// TIA Portal project "Industry 4.0_Plant_Logic" (V16)

(* hardware
DEVICE "S7-1200 station_1"  S7-1200 Station
   slot 0: "Rack_0"  S7-1200 Rack  Rack  V1.0
   slot 1: "S7_1212"  CPU 1212C AC/DC/Rly  6ES7 212-1BE40-0XB0  V4.4
   slot 2: "AQ 2x14BIT_1"  SM 1232 AQ2  6ES7 232-4HB32-0XB0  V2.1
DEVICE "HMI_1"  KTP700 Basic PN
   slot 0: "HMI_1"  KTP700 Basic PN  6AV2 123-2GB03-0AX0  15.1.0.0
   slot 1: "HMI_RT_1"  KTP700 Basic PN  6AV2 123-2GB03-0AX0  15.1.0.0
   slot 5: "HMI_1.IE_CP_1"  PROFINET Interface  15.0.1.0
      slot 1: "PROFINET Interface_1"  PROFINET Interface
         slot 1: "Port_1"  Port
*)

// ===== PLC "S7_1212"  CPU 1212C AC/DC/Rly =====

VAR_GLOBAL   // PLC tag table "Default tag table"
   "FIC_B102" AT %IW64 : Int;   // Flow meter(0 - 27648)
   "LIC_B101" AT %IW66 : Int;   // Tank02 Level meter(0 - 27648)
   "PS1_RFID_Station" AT %I0.0 : Bool;   // PS-Proximity Switch
   "PS2_Filling_Station" AT %I0.1 : Bool;
   "PS3_Quality_Station" AT %I0.2 : Bool;
   "PS4_End_of_Conveyor" AT %I0.3 : Bool;
   "T01_Low_Level" AT %I0.4 : Bool;   // Proximity sensor measuring Low level of Tank01
   "T01_High_Level" AT %I0.5 : Bool;   // Proximity sensor measuring High level of Tank01
   "T01_Outlet" AT %Q0.1 : Bool;   // Tank01 Output Solenoid Valve
   "T02_Outlet" AT %Q0.2 : Bool;   // Tank02 Output Solenoid Valve
   "Outlet_Pump_Motor" AT %Q0.3 : Bool;   // Pump Motor
   "Conveyor_Motor" AT %Q0.0 : Bool;
   "NTRG_06" AT %M5.5 : Bool;
   "NTRG_09" AT %M5.6 : Bool;
   "NTRG_099" AT %M5.7 : Bool;
   "PTRG10" AT %M6.0 : Bool;
   "PTRIG999" AT %M6.1 : Bool;
   "PTRIG998" AT %M6.2 : Bool;
   "PTRIG888" AT %M6.3 : Bool;
   "ptrig141" AT %M6.4 : Bool;
   "ptrig142" AT %M6.5 : Bool;
   "ptrig143" AT %M6.6 : Bool;
   "Ptrig241" AT %M6.7 : Bool;
   "reset__bottle_animation_timer" AT %M7.0 : Bool;
   "motor_running_time" AT %MD8 : Time;
   "ntrig555" AT %M7.1 : Bool;
   "Total Bottle filled" AT %MW8 : Int;
   "abc" AT %QW98 : Int;
   "Static_1" AT %MW12 : Int;
   "Static_1(1)" AT %MW14 : Int;
   "Static_1(2)" AT %MW16 : Int;
   "i" AT %MW18 : Int;
   "ONS_1" AT %M7.2 : Bool;
END_VAR

VAR_GLOBAL   // PLC tag table "P_N_TRIG"
   "PTRIG1" AT %M0.0 : Bool;
   "PTRIG2" AT %M0.1 : Bool;
   "PTRIG3" AT %M0.2 : Bool;
   "PTRIG4" AT %M0.3 : Bool;
   "PTRIG5" AT %M0.4 : Bool;
   "PTRIG6" AT %M0.5 : Bool;
   "PTRIG7" AT %M0.6 : Bool;
   "PTRIG8" AT %M0.7 : Bool;
   "PTRIG9" AT %M1.0 : Bool;
   "PTRIG10" AT %M1.1 : Bool;
   "PTRIG11" AT %M1.2 : Bool;
   "PTRIG12" AT %M1.3 : Bool;
   "PTRIG13" AT %M1.4 : Bool;
   "PTRIG14" AT %M1.5 : Bool;
   "PTRIG15" AT %M1.6 : Bool;
   "PTRIG16" AT %M1.7 : Bool;
   "PTRIG17" AT %M2.0 : Bool;
   "PTRIG18" AT %M2.1 : Bool;
   "PTRIG19" AT %M2.2 : Bool;
   "PTRIG20" AT %M2.3 : Bool;
   "PTRIG21" AT %M2.4 : Bool;
   "PTRIG22" AT %M2.5 : Bool;
   "PTRIG23" AT %M2.6 : Bool;
   "NTRIG1" AT %M2.7 : Bool;
   "NTRIG2" AT %M3.0 : Bool;
   "NTRIG3" AT %M3.1 : Bool;
   "NTRIG4" AT %M3.2 : Bool;
   "NTRIG5" AT %M3.3 : Bool;
   "NTRIG6" AT %M3.4 : Bool;
   "NTRIG7" AT %M3.5 : Bool;
   "NTRIG8" AT %M3.6 : Bool;
   "NTRIG9" AT %M3.7 : Bool;
   "NTRIG10" AT %M4.0 : Bool;
   "NTRIG11" AT %M4.1 : Bool;
   "NTRIG12" AT %M4.2 : Bool;
   "NTRIG13" AT %M4.3 : Bool;
   "NTRIG14" AT %M4.4 : Bool;
   "NTRIG15" AT %M4.5 : Bool;
   "NTRIG16" AT %M4.6 : Bool;
   "NTRIG17" AT %M4.7 : Bool;
   "NTRIG18" AT %M5.0 : Bool;
   "NTRIG19" AT %M5.1 : Bool;
   "NTRIG20" AT %M5.2 : Bool;
   "PTRIG24" AT %M5.3 : Bool;
   "PTRIG25" AT %M5.4 : Bool;
END_VAR

DATA_BLOCK "Global_DB"   // DB1
{ S7_Optimized_Access := 'TRUE' }
VERSION : 0.1
   VAR
      Input : Struct   // Values from input devices
         FIC_B102 : Int;   // Flow in (0-27648) range
         LIC_B101 : Int;   // Level in (0-27648) range
         PS1_RFID_Station : Bool;   // Proximity sensor at RFID station
         PS2_Filling_Station : Bool;   // Proximity sensor at Filling station
         PS3_Quality_Station : Bool;   // Proximity sensor at Quality Station
         PS4_End_of_Conveyor : Bool;   // Proximity sensor at End of the conveyor
         T01_Low_Level : Bool;   // Tank01 Low level detection sensor
         T01_High_Level : Bool;   // Tank01 High level detection sensor
      END_STRUCT;
      Output : Struct   // Values to Output devices
         T01_Outlet : Bool;   // Tank01 Outlet Solenoid Valve
         T02_Outlet : Bool;   // Tank02 Outlet Solenoid Valve
         Outlet_Pump_Motor : Bool;   // To tigger Pump motor relay
         Conveyor_Motor : Bool;   // To tigger Conveyor motor relay
         T01_Inlet : Bool;   // Tank01 Inlet Solenoid Valve(Not implemented)
         T02_Inlet : Bool;   // Tank02 Inlet Solenoid Valve(Not implemented)
      END_STRUCT;
      Other_Parameters : Struct   // Scalled and middle Variables
         Liquid_A_Filled : Bool;   // Liquid_A_filled flag activated when intended amount of Liquid A is filled
         Add_Done : Bool;
         Liquid_B_Filled : Bool;   // Liquid_B_filled flag activated when intended amount of Liquid B is filled
         Flow_ml_per_sec : Real;   // Scalled flow meter reading (0-250mL/sec)
         LiquidA_in_Bottle_ml : Real;
         LiquidB_in_Bottle_ml : Real;
         T02_Level_in_L : Real;   // Scalled level meter reading (0-10L)
         T02_High_Level_Limit : Real;
         T02_Low_Level_Limit : Real;
         Alarm_Reset : Bool;   // to reset all active alarms
         operation_cycle_time : Time;   // Time taken for the filling of one bottle
         index : Int := 1;
      END_STRUCT;
      Error : Struct
         Alarm : Word;
      END_STRUCT;
      Master_Commands : Struct
         operation_finished : Bool;
         operation_begin : Bool;
         Order_Variables : Struct   // Online Order parameter
            "Total Bottle filled" : Int;
            Order_ID : UInt;
            Quantity : UInt := 0;   // Quanity of bottle to be filled in pesent order
            Liquid_A_pct : Int := 0;   // data from RFID tags or Order
            Liquid_B_pct : Int;   // datafrom RFID tags or Order
            Order_received : Bool;   // Activated when new order is received.
            Bottle_Count : Int := 1;   // Total Bottle filled
            Order_completed : Bool;   // Order completion flag(After filling all bottle)
         END_STRUCT;
      END_STRUCT;
      SCADA : Struct   // SCADA animation tags
         motor_running_time : Time;   // To display bottle moving on the conveyor based on the running time of conveyor
      END_STRUCT;
      Flow : Real;
      Motor_Output_PCT : Int;
      Production_Data : Struct   // Unit ml
         Total_Liquid_in_Bottle : Array[1..5] of Real;
         LiquidA_in_Bottle : Array[1..5] of Real;
         operation_cycles : Array[1..5] of Time;
         LiquidB_in_Bottle : Array[1..5] of Real;
         current_cycle : Int := 1;
      END_STRUCT;
      Array_Voltage : Array[0..999] of Real;
      Voltage_Timer : Bool;
      "Locking bits" : Struct
         Starting_station_bit : Bool;
         Filling_station_bit : Bool;
         Quality_station_bit : Bool;
         End_station_bit : Bool;
      END_STRUCT;
   END_VAR
BEGIN
END_DATA_BLOCK

// folder: Function Blocks

DATA_BLOCK "Re-filling_Logic_DB"   // DB2
{ S7_Optimized_Access := 'TRUE' }
VERSION : 0.1
// stored: InstanceOfName Re-filling_Logic
"Re-filling_Logic"
BEGIN
END_DATA_BLOCK

DATA_BLOCK "Filling_Logic_DB"   // DB4
{ S7_Optimized_Access := 'TRUE' }
VERSION : 0.1
// stored: InstanceOfName Filling_Logic
"Filling_Logic"
BEGIN
END_DATA_BLOCK

DATA_BLOCK "Filling_Logic_DB_1"   // DB5
{ S7_Optimized_Access := 'TRUE' }
VERSION : 0.1
// stored: InstanceOfName Filling_Logic
"Filling_Logic"
BEGIN
END_DATA_BLOCK

DATA_BLOCK "Alarm_Logic_DB"   // DB7
{ S7_Optimized_Access := 'TRUE' }
VERSION : 0.1
// stored: InstanceOfName Alarm_Logic
"Alarm_Logic"
BEGIN
END_DATA_BLOCK

DATA_BLOCK "Tank1_DB"   // DB9
{ S7_Optimized_Access := 'TRUE' }
VERSION : 0.1
// stored: InstanceOfName Tank1
"Tank1"
BEGIN
END_DATA_BLOCK

DATA_BLOCK "Tank2_DB"   // DB10
{ S7_Optimized_Access := 'TRUE' }
VERSION : 0.1
// stored: InstanceOfName Tank2
"Tank2"
BEGIN
END_DATA_BLOCK

DATA_BLOCK "ProductionData_Reset_DB"   // DB13
{ S7_Optimized_Access := 'TRUE' }
VERSION : 0.1
// stored: InstanceOfName ProductionData_Reset
"ProductionData_Reset"
BEGIN
END_DATA_BLOCK

DATA_BLOCK "Operation_cycle_DB"   // DB15
{ S7_Optimized_Access := 'TRUE' }
VERSION : 0.1
// stored: InstanceOfName Operation_cycle
"Operation_cycle"
BEGIN
END_DATA_BLOCK

DATA_BLOCK "Reseting_order_DB"   // DB18
{ S7_Optimized_Access := 'TRUE' }
VERSION : 0.1
// stored: InstanceOfName Reseting_order
"Reseting_order"
BEGIN
END_DATA_BLOCK

DATA_BLOCK "Array_Voltage_Logic_DB_1"   // DB25
{ S7_Optimized_Access := 'TRUE' }
VERSION : 0.1
// stored: InstanceOfName Array_Voltage_Logic
"Array_Voltage_Logic"
BEGIN
END_DATA_BLOCK

// folder: System blocks/Program resources

DATA_BLOCK "IEC_Timer_6_DB_1"   // DB3
{ S7_Optimized_Access := 'TRUE' }
AUTHOR : Simatic
FAMILY : IEC
NAME : IEC_TMR
VERSION : 1.0
// stored: InstanceOfName IEC_TIMER
"IEC_TIMER"
BEGIN
END_DATA_BLOCK

DATA_BLOCK "IEC_Timer_0_DB_1"   // DB6
{ S7_Optimized_Access := 'TRUE' }
AUTHOR : Simatic
FAMILY : IEC
NAME : IEC_TMR
VERSION : 1.0
// stored: InstanceOfName IEC_TIMER
"IEC_TIMER"
BEGIN
END_DATA_BLOCK

DATA_BLOCK "IEC_Timer_0_DB_999"   // DB8
{ S7_Optimized_Access := 'TRUE' }
AUTHOR : Simatic
FAMILY : IEC
NAME : IEC_TMR
VERSION : 1.0
// stored: InstanceOfName IEC_TIMER
"IEC_TIMER"
BEGIN
END_DATA_BLOCK

DATA_BLOCK "IEC_Timer_0_DB_7"   // DB11
{ S7_Optimized_Access := 'TRUE' }
AUTHOR : Simatic
FAMILY : IEC
NAME : IEC_TMR
VERSION : 1.0
// stored: InstanceOfName IEC_TIMER
"IEC_TIMER"
BEGIN
END_DATA_BLOCK

DATA_BLOCK "IEC_Counter_0_DB"   // DB12
{ S7_Optimized_Access := 'TRUE' }
AUTHOR : Simatic
FAMILY : IEC
NAME : CNTR
VERSION : 1.0
// stored: InstanceOfName IEC_COUNTER
"IEC_COUNTER"
BEGIN
END_DATA_BLOCK

DATA_BLOCK "Cycle_time"   // DB14
{ S7_Optimized_Access := 'TRUE' }
AUTHOR : Simatic
FAMILY : IEC
NAME : IEC_TMR
VERSION : 1.0
// stored: InstanceOfName IEC_TIMER
"IEC_TIMER"
BEGIN
END_DATA_BLOCK

DATA_BLOCK "IEC_Timer_655"   // DB16
{ S7_Optimized_Access := 'TRUE' }
AUTHOR : Simatic
FAMILY : IEC
NAME : IEC_TMR
VERSION : 1.0
// stored: InstanceOfName IEC_TIMER
"IEC_TIMER"
BEGIN
END_DATA_BLOCK

DATA_BLOCK "Waiting time"   // DB20
{ S7_Optimized_Access := 'TRUE' }
AUTHOR : Simatic
FAMILY : IEC
NAME : IEC_TMR
VERSION : 1.0
// stored: InstanceOfName IEC_TIMER
"IEC_TIMER"
BEGIN
END_DATA_BLOCK

// folder: (top level)

ORGANIZATION_BLOCK "Main"   // OB1, LAD, ProgramCycle
TITLE = "Main Program Sweep (Cycle)"
{ S7_Optimized_Access := 'TRUE' }
VERSION : 0.1
   VAR_INPUT
      Initial_Call : Bool;   // Initial call of this OB
      Remanence : Bool;   // =True, if remanent data are available
   END_VAR
   VAR_TEMP   // added for the SCL form of the ladder/FBD networks
      _w1 : Bool;
      _w2 : Bool;
   END_VAR
BEGIN

REGION Network 1: Tank 1 and Tank 2 re-filling Logic
   // 1."Re-filling_logic" block is logic block to refill liquid in tanks based on their levels(Hardware not present yet)
   // 2."Operation_cycle" block to measure the time of bottle filling which starts from picking bottle till bottle placed.
   // 3."Reading" Mapping from Physical address to Global_DB (for input devices)
   // 4."Writing" Mapping from Global_DB to Physical address(for output devices)
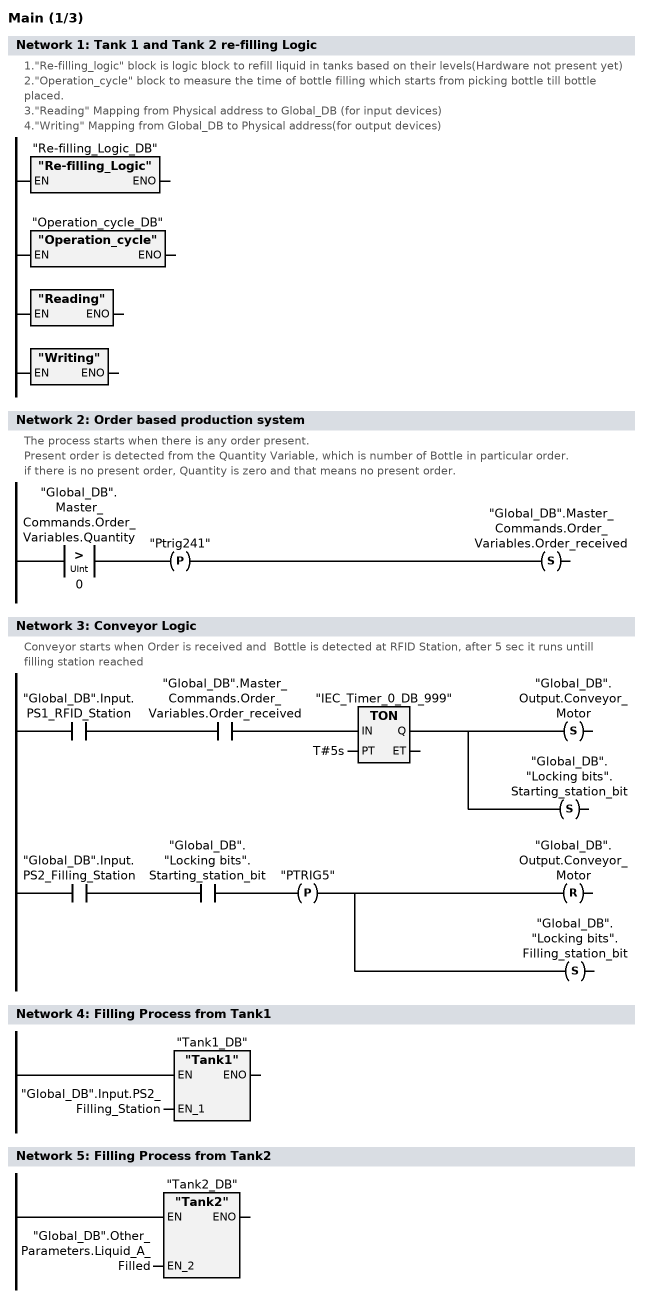
   RUNG wire#powerrail
      "Re-filling_Logic_DB"()
   END_RUNG
   RUNG wire#powerrail
      "Operation_cycle_DB"()
   END_RUNG
   RUNG wire#powerrail
      "Reading"()
   END_RUNG
   RUNG wire#powerrail
      "Writing"()
   END_RUNG
   // the same network as SCL:
   "Re-filling_Logic_DB"();   // "Re-filling_Logic"
   "Operation_cycle_DB"();   // "Operation_cycle"
   "Reading"();
   "Writing"();
END_REGION

REGION Network 2: Order based production system
   // The process starts when there is any order present.
   // Present order is detected from the Quantity Variable, which is number of Bottle in particular order.
   // if there is no present order, Quantity is zero and that means no present order.
   RUNG wire#powerrail
      { S7_Templates := "SrcType := UInt" } GT_Contact(in1 := "Global_DB".Master_Commands.Order_Variables.Quantity, in2 := 0)
      P_Trig( "Ptrig241" )
      S_Coil( "Global_DB".Master_Commands.Order_Variables.Order_received )
   END_RUNG
   // the same network as SCL:
   #_w1 := "Global_DB".Master_Commands.Order_Variables.Quantity > 0;
   #_w2 := #_w1 AND NOT "Ptrig241";   // rising edge
   "Ptrig241" := #_w1;
   IF #_w2 THEN "Global_DB".Master_Commands.Order_Variables.Order_received := TRUE; END_IF;
END_REGION

REGION Network 3: Conveyor Logic
   // Conveyor starts when Order is received and  Bottle is detected at RFID Station, after 5 sec it runs untill filling station reached
   "IEC_Timer_0_DB_999".TON(IN := "Global_DB".Input.PS1_RFID_Station AND "Global_DB".Master_Commands.Order_Variables.Order_received,
                           PT := T#5s);
   IF "IEC_Timer_0_DB_999".Q THEN
       "Global_DB".Output.Conveyor_Motor := TRUE;
       "Global_DB"."Locking bits".Starting_station_bit := TRUE;
   END_IF;
   #_w1 := "Global_DB".Input.PS2_Filling_Station AND "Global_DB"."Locking bits".Starting_station_bit;
   #_w2 := #_w1 AND NOT "PTRIG5";   // rising edge
   "PTRIG5" := #_w1;
   IF #_w2 THEN
       "Global_DB".Output.Conveyor_Motor := FALSE;
       "Global_DB"."Locking bits".Filling_station_bit := TRUE;
   END_IF;
END_REGION

REGION Network 4: Filling Process from Tank1
   RUNG wire#powerrail
      "Tank1_DB"(EN_1 := "Global_DB".Input.PS2_Filling_Station)
   END_RUNG
   // the same network as SCL:
   "Tank1_DB"(EN_1 := "Global_DB".Input.PS2_Filling_Station);   // "Tank1"
END_REGION

REGION Network 5: Filling Process from Tank2
   RUNG wire#powerrail
      "Tank2_DB"(EN_2 := "Global_DB".Other_Parameters.Liquid_A_Filled)
   END_RUNG
   // the same network as SCL:
   "Tank2_DB"(EN_2 := "Global_DB".Other_Parameters.Liquid_A_Filled);   // "Tank2"
END_REGION

REGION Network 6: Store data in database for records
   // after filling the liquid from both tanks, ADD block adds the value of filled amount of Liquid A nad Liquid B in the bottle to keep record of total liquid filled in particular bottle.
   // 
   // then bottle number is incremented.
   // 
   // Values reset for next cycle.
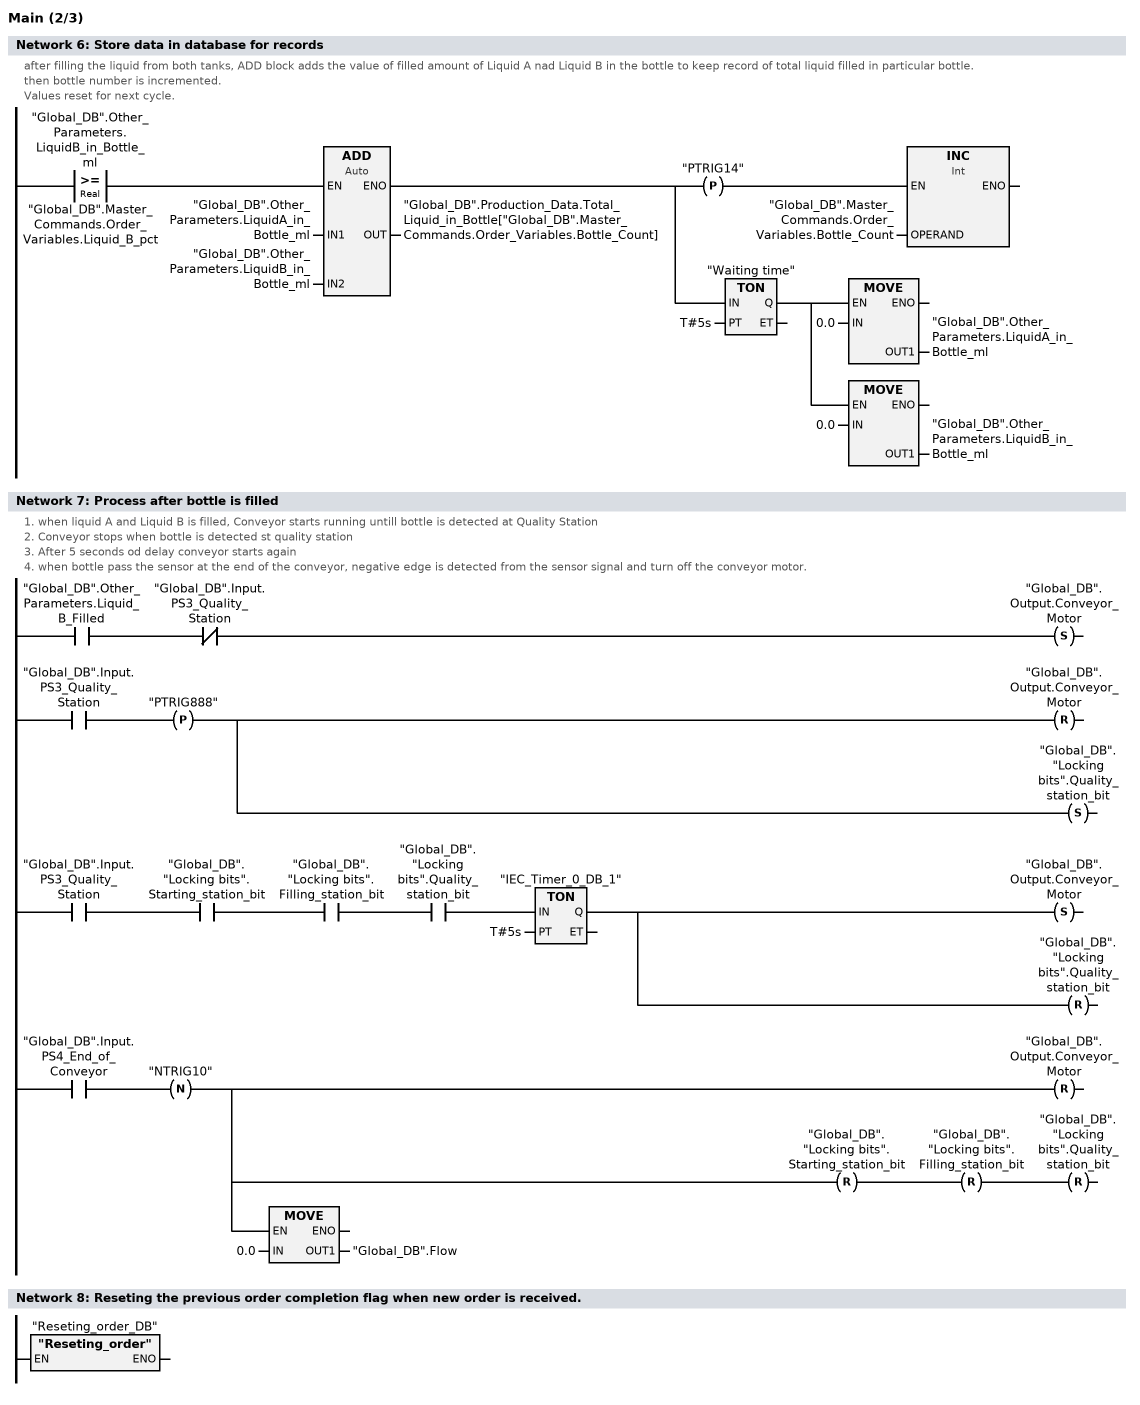
   #_w1 := "Global_DB".Other_Parameters.LiquidB_in_Bottle_ml >= "Global_DB".Master_Commands.Order_Variables.Liquid_B_pct;
   IF #_w1 THEN
       "Global_DB".Production_Data.Total_Liquid_in_Bottle["Global_DB".Master_Commands.Order_Variables.Bottle_Count] := "Global_DB".Other_Parameters.LiquidA_in_Bottle_ml + "Global_DB".Other_Parameters.LiquidB_in_Bottle_ml;
   END_IF;
   #_w2 := #_w1 AND NOT "PTRIG14";   // rising edge
   "PTRIG14" := #_w1;
   IF #_w2 THEN
       "Global_DB".Master_Commands.Order_Variables.Bottle_Count := "Global_DB".Master_Commands.Order_Variables.Bottle_Count + 1;
   END_IF;
   "Waiting time".TON(IN := #_w1, PT := T#5s);
   IF "Waiting time".Q THEN
       "Global_DB".Other_Parameters.LiquidA_in_Bottle_ml := 0.0;
       "Global_DB".Other_Parameters.LiquidB_in_Bottle_ml := 0.0;
   END_IF;
END_REGION

REGION Network 7: Process after bottle is filled
   // 1. when liquid A and Liquid B is filled, Conveyor starts running untill bottle is detected at Quality Station
   // 2. Conveyor stops when bottle is detected st quality station
   // 3. After 5 seconds od delay conveyor starts again
   // 4. when bottle pass the sensor at the end of the conveyor, negative edge is detected from the sensor signal and turn off the conveyor motor.
   IF "Global_DB".Other_Parameters.Liquid_B_Filled AND NOT "Global_DB".Input.PS3_Quality_Station THEN
       "Global_DB".Output.Conveyor_Motor := TRUE;
   END_IF;
   #_w1 := "Global_DB".Input.PS3_Quality_Station AND NOT "PTRIG888";   // rising edge
   "PTRIG888" := "Global_DB".Input.PS3_Quality_Station;
   IF #_w1 THEN
       "Global_DB".Output.Conveyor_Motor := FALSE;
       "Global_DB"."Locking bits".Quality_station_bit := TRUE;
   END_IF;
   "IEC_Timer_0_DB_1".TON(IN := "Global_DB".Input.PS3_Quality_Station AND "Global_DB"."Locking bits".Starting_station_bit AND "Global_DB"."Locking bits".Filling_station_bit AND "Global_DB"."Locking bits".Quality_station_bit,
                          PT := T#5s);
   IF "IEC_Timer_0_DB_1".Q THEN
       "Global_DB".Output.Conveyor_Motor := TRUE;
       "Global_DB"."Locking bits".Quality_station_bit := FALSE;
   END_IF;
   #_w2 := NOT "Global_DB".Input.PS4_End_of_Conveyor AND "NTRIG10";   // falling edge
   "NTRIG10" := "Global_DB".Input.PS4_End_of_Conveyor;
   IF #_w2 THEN
       "Global_DB".Output.Conveyor_Motor := FALSE;
       "Global_DB"."Locking bits".Starting_station_bit := FALSE;
       "Global_DB"."Locking bits".Filling_station_bit := FALSE;
       "Global_DB"."Locking bits".Quality_station_bit := FALSE;
       "Global_DB".Flow := 0.0;
   END_IF;
END_REGION

REGION Network 8: Reseting the previous order completion flag when new order is received.
   RUNG wire#powerrail
      "Reseting_order_DB"()
   END_RUNG
   // the same network as SCL:
   "Reseting_order_DB"();   // "Reseting_order"
END_REGION

REGION Network 9: Reseting Production data after each order completion
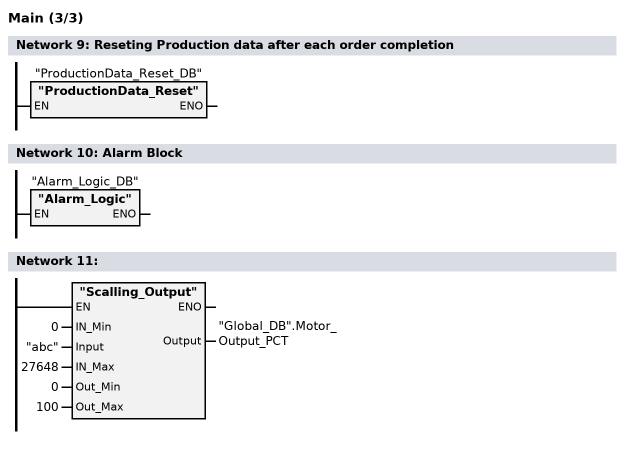
   RUNG wire#powerrail
      "ProductionData_Reset_DB"()
   END_RUNG
   // the same network as SCL:
   "ProductionData_Reset_DB"();   // "ProductionData_Reset"
END_REGION

REGION Network 10: Alarm Block
   RUNG wire#powerrail
      "Alarm_Logic_DB"()
   END_RUNG
   // the same network as SCL:
   "Alarm_Logic_DB"();   // "Alarm_Logic"
END_REGION

REGION Network 11
   RUNG wire#powerrail
      "Scalling_Output"(IN_Min := 0, Input := "abc", IN_Max := 27648, Out_Min := 0, Out_Max := 100, Output => "Global_DB".Motor_Output_PCT)
   END_RUNG
   // the same network as SCL:
   "Scalling_Output"(IN_Min := 0,
                     Input := "abc",
                     IN_Max := 27648,
                     Out_Min := 0,
                     Out_Max := 100,
                     Output => "Global_DB".Motor_Output_PCT);
END_REGION
END_ORGANIZATION_BLOCK

ORGANIZATION_BLOCK "Totalizer"   // OB30, LAD, CyclicInterrupt
TITLE = This Totalizer [OB30] block runs every 1 second
{ S7_Optimized_Access := 'TRUE' }
VERSION : 0.1
// This block is programmed to get quantity of liquid (ml) which passed from flow meter(mL\sec).
// 
// By adding flow meter reading at every second, we can quantity of liquid for specific time.
   VAR_INPUT
      Initial_Call : Bool;   // Initial call of this OB
      Event_Count : Int;   // Events discarded
   END_VAR
BEGIN

REGION Network 1: Tank1 - LiquidA filling value Totalizer
   // 1. When tank01 outlet valve is opened, means process of Liquid A is filling in the Bottle.
   // 
   // By addting flow meter reading every one second, how much liquid A is filled in the bottle is calculated.
   // 
   // 2. When amount of liquidA exceeds than what we want to fill in the particular bottle, "Liquid_A_Filled" flag is activated and Tank01 outlet valve is closed.
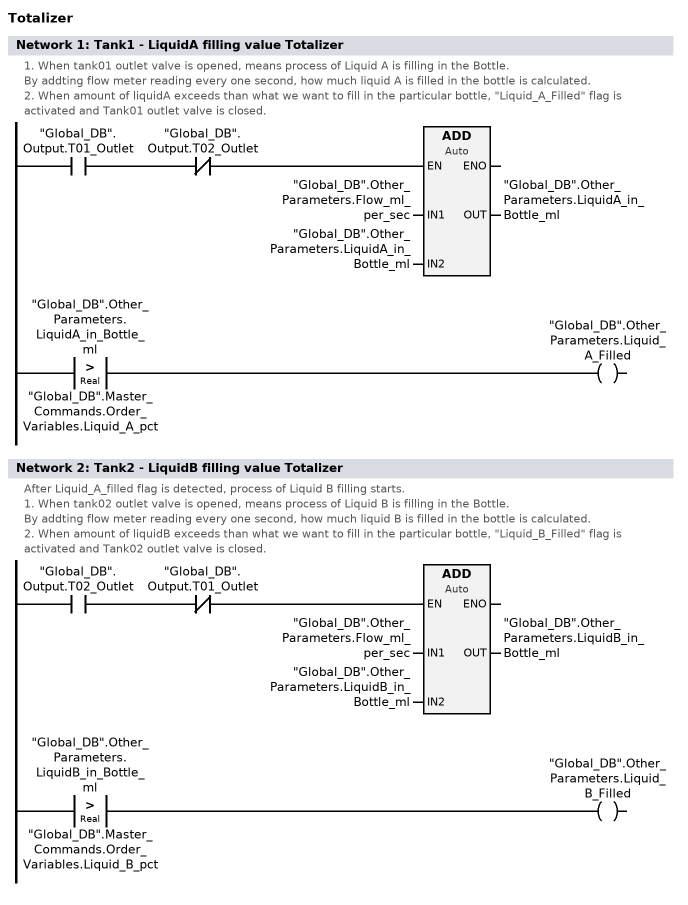
   RUNG wire#powerrail
      Contact( "Global_DB".Output.T01_Outlet )
      I_Contact( "Global_DB".Output.T02_Outlet )
      Add(in1 := "Global_DB".Other_Parameters.Flow_ml_per_sec, in2 := "Global_DB".Other_Parameters.LiquidA_in_Bottle_ml, out => "Global_DB".Other_Parameters.LiquidA_in_Bottle_ml)
   END_RUNG
   RUNG wire#powerrail
      { S7_Templates := "SrcType := Real" } GT_Contact(in1 := "Global_DB".Other_Parameters.LiquidA_in_Bottle_ml, in2 := "Global_DB".Master_Commands.Order_Variables.Liquid_A_pct)
      Coil( "Global_DB".Other_Parameters.Liquid_A_Filled )
   END_RUNG
   // the same network as SCL:
   IF "Global_DB".Output.T01_Outlet AND NOT "Global_DB".Output.T02_Outlet THEN
       "Global_DB".Other_Parameters.LiquidA_in_Bottle_ml := "Global_DB".Other_Parameters.Flow_ml_per_sec + "Global_DB".Other_Parameters.LiquidA_in_Bottle_ml;
   END_IF;
   "Global_DB".Other_Parameters.Liquid_A_Filled := "Global_DB".Other_Parameters.LiquidA_in_Bottle_ml > "Global_DB".Master_Commands.Order_Variables.Liquid_A_pct;
END_REGION

REGION Network 2: Tank2 - LiquidB filling value Totalizer
   // After Liquid_A_filled flag is detected, process of Liquid B filling starts.
   // 
   // 1. When tank02 outlet valve is opened, means process of Liquid B is filling in the Bottle.
   // 
   // By addting flow meter reading every one second, how much liquid B is filled in the bottle is calculated.
   // 
   // 2. When amount of liquidB exceeds than what we want to fill in the particular bottle, "Liquid_B_Filled" flag is activated and Tank02 outlet valve is closed.
   RUNG wire#powerrail
      Contact( "Global_DB".Output.T02_Outlet )
      I_Contact( "Global_DB".Output.T01_Outlet )
      Add(in1 := "Global_DB".Other_Parameters.Flow_ml_per_sec, in2 := "Global_DB".Other_Parameters.LiquidB_in_Bottle_ml, out => "Global_DB".Other_Parameters.LiquidB_in_Bottle_ml)
   END_RUNG
   RUNG wire#powerrail
      { S7_Templates := "SrcType := Real" } GT_Contact(in1 := "Global_DB".Other_Parameters.LiquidB_in_Bottle_ml, in2 := "Global_DB".Master_Commands.Order_Variables.Liquid_B_pct)
      Coil( "Global_DB".Other_Parameters.Liquid_B_Filled )
   END_RUNG
   // the same network as SCL:
   IF "Global_DB".Output.T02_Outlet AND NOT "Global_DB".Output.T01_Outlet THEN
       "Global_DB".Other_Parameters.LiquidB_in_Bottle_ml := "Global_DB".Other_Parameters.Flow_ml_per_sec + "Global_DB".Other_Parameters.LiquidB_in_Bottle_ml;
   END_IF;
   "Global_DB".Other_Parameters.Liquid_B_Filled := "Global_DB".Other_Parameters.LiquidB_in_Bottle_ml > "Global_DB".Master_Commands.Order_Variables.Liquid_B_pct;
END_REGION
END_ORGANIZATION_BLOCK

ORGANIZATION_BLOCK "Cyclic interrupt"   // OB31, LAD, CyclicInterrupt
{ S7_Optimized_Access := 'TRUE' }
VERSION : 0.1
   VAR_INPUT
      Initial_Call : Bool;   // Initial call of this OB
      Event_Count : Int;   // Events discarded
   END_VAR
   VAR_TEMP
      TV_A : Real;
      TV_B : Real;
   END_VAR
BEGIN

REGION Network 1
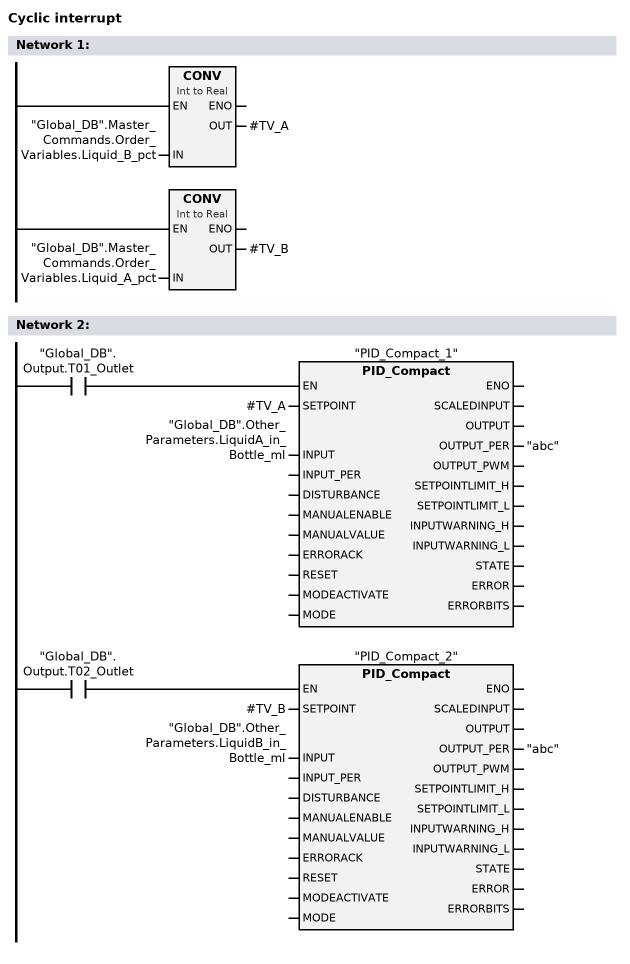
   RUNG wire#powerrail
      { S7_Templates := "[SrcType := Int, DestType := Real]" } Convert(in := "Global_DB".Master_Commands.Order_Variables.Liquid_B_pct, out => #TV_A)
   END_RUNG
   RUNG wire#powerrail
      { S7_Templates := "[SrcType := Int, DestType := Real]" } Convert(in := "Global_DB".Master_Commands.Order_Variables.Liquid_A_pct, out => #TV_B)
   END_RUNG
   // the same network as SCL:
   #TV_A := INT_TO_REAL("Global_DB".Master_Commands.Order_Variables.Liquid_B_pct);
   #TV_B := INT_TO_REAL("Global_DB".Master_Commands.Order_Variables.Liquid_A_pct);
END_REGION

REGION Network 2
   IF "Global_DB".Output.T01_Outlet THEN
       "PID_Compact_1"(Setpoint := #TV_A,   // PID_Compact
                       Input := "Global_DB".Other_Parameters.LiquidA_in_Bottle_ml,
                       Output_PER => "abc");
   END_IF;
   IF "Global_DB".Output.T02_Outlet THEN
       "PID_Compact_2"(Setpoint := #TV_B,   // PID_Compact
                       Input := "Global_DB".Other_Parameters.LiquidB_in_Bottle_ml,
                       Output_PER => "abc");
   END_IF;
END_REGION
END_ORGANIZATION_BLOCK

ORGANIZATION_BLOCK "Total flow calculator"   // OB32, SCL, CyclicInterrupt
{ S7_Optimized_Access := 'TRUE' }
VERSION : 0.1
   VAR_INPUT
      Initial_Call : Bool;   // Initial call of this OB
      Event_Count : Int;   // Events discarded
   END_VAR
BEGIN
   IF "Outlet_Pump_Motor" = TRUE THEN

       "Global_DB".Flow := "Global_DB".Flow + "Global_DB".Other_Parameters.Flow_ml_per_sec;

   END_IF;
END_ORGANIZATION_BLOCK

ORGANIZATION_BLOCK "Voltage"   // OB33, LAD, CyclicInterrupt
{ S7_Optimized_Access := 'TRUE' }
VERSION : 0.1
   VAR_INPUT
      Initial_Call : Bool;   // Initial call of this OB
      Event_Count : Int;   // Events discarded
   END_VAR
BEGIN

REGION Network 1
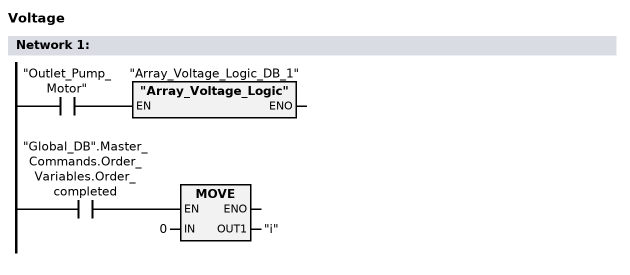
   RUNG wire#powerrail
      Contact( "Outlet_Pump_Motor" )
      "Array_Voltage_Logic_DB_1"()
   END_RUNG
   RUNG wire#powerrail
      Contact( "Global_DB".Master_Commands.Order_Variables.Order_completed )
      Move(in := 0, out1 => "i")
   END_RUNG
   // the same network as SCL:
   IF "Outlet_Pump_Motor" THEN
       "Array_Voltage_Logic_DB_1"();   // "Array_Voltage_Logic"
   END_IF;
   IF "Global_DB".Master_Commands.Order_Variables.Order_completed THEN "i" := 0; END_IF;
END_REGION
END_ORGANIZATION_BLOCK

// folder: Function Blocks

FUNCTION_BLOCK "Re-filling_Logic"   // FB1, LAD
{ S7_Optimized_Access := 'TRUE' }
VERSION : 0.1
   VAR_TEMP   // added for the SCL form of the ladder/FBD networks
      _w1 : Bool;
      _w2 : Bool;
      _w3 : Bool;
      _w4 : Bool;
   END_VAR
BEGIN

REGION Network 1: Tank2 Re-filling Proccess
   // When liquid level in Tank02 is below low limit, T02 inlet valve is opened till level reached at high limit.
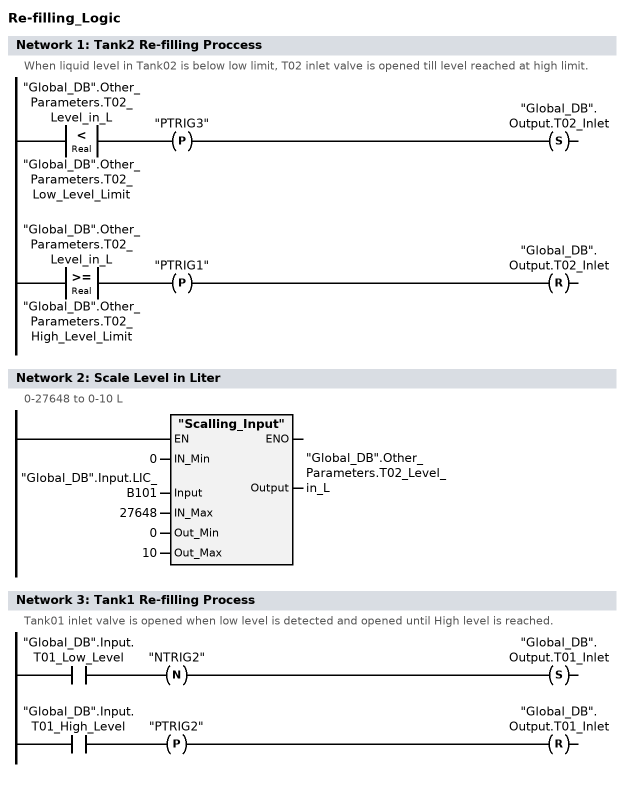
   RUNG wire#powerrail
      { S7_Templates := "SrcType := Real" } LT_Contact(in1 := "Global_DB".Other_Parameters.T02_Level_in_L, in2 := "Global_DB".Other_Parameters.T02_Low_Level_Limit)
      P_Trig( "PTRIG3" )
      S_Coil( "Global_DB".Output.T02_Inlet )
   END_RUNG
   RUNG wire#powerrail
      { S7_Templates := "SrcType := Real" } GE_Contact(in1 := "Global_DB".Other_Parameters.T02_Level_in_L, in2 := "Global_DB".Other_Parameters.T02_High_Level_Limit)
      P_Trig( "PTRIG1" )
      R_Coil( "Global_DB".Output.T02_Inlet )
   END_RUNG
   // the same network as SCL:
   #_w1 := "Global_DB".Other_Parameters.T02_Level_in_L < "Global_DB".Other_Parameters.T02_Low_Level_Limit;
   #_w2 := #_w1 AND NOT "PTRIG3";   // rising edge
   "PTRIG3" := #_w1;
   IF #_w2 THEN "Global_DB".Output.T02_Inlet := TRUE; END_IF;
   #_w3 := "Global_DB".Other_Parameters.T02_Level_in_L >= "Global_DB".Other_Parameters.T02_High_Level_Limit;
   #_w4 := #_w3 AND NOT "PTRIG1";   // rising edge
   "PTRIG1" := #_w3;
   IF #_w4 THEN "Global_DB".Output.T02_Inlet := FALSE; END_IF;
END_REGION

REGION Network 2: Scale Level in Liter
   // 0-27648 to 0-10 L
   RUNG wire#powerrail
      "Scalling_Input"(IN_Min := 0, Input := "Global_DB".Input.LIC_B101, IN_Max := 27648, Out_Min := 0, Out_Max := 10, Output => "Global_DB".Other_Parameters.T02_Level_in_L)
   END_RUNG
   // the same network as SCL:
   "Scalling_Input"(IN_Min := 0,
                    Input := "Global_DB".Input.LIC_B101,
                    IN_Max := 27648,
                    Out_Min := 0,
                    Out_Max := 10,
                    Output => "Global_DB".Other_Parameters.T02_Level_in_L);
END_REGION

REGION Network 3: Tank1 Re-filling Process
   // Tank01 inlet valve is opened when low level is detected and opened until High level is reached.
   RUNG wire#powerrail
      Contact( "Global_DB".Input.T01_Low_Level )
      N_Trig( "NTRIG2" )
      S_Coil( "Global_DB".Output.T01_Inlet )
   END_RUNG
   RUNG wire#powerrail
      Contact( "Global_DB".Input.T01_High_Level )
      P_Trig( "PTRIG2" )
      R_Coil( "Global_DB".Output.T01_Inlet )
   END_RUNG
   // the same network as SCL:
   #_w1 := NOT "Global_DB".Input.T01_Low_Level AND "NTRIG2";   // falling edge
   "NTRIG2" := "Global_DB".Input.T01_Low_Level;
   IF #_w1 THEN "Global_DB".Output.T01_Inlet := TRUE; END_IF;
   #_w2 := "Global_DB".Input.T01_High_Level AND NOT "PTRIG2";   // rising edge
   "PTRIG2" := "Global_DB".Input.T01_High_Level;
   IF #_w2 THEN "Global_DB".Output.T01_Inlet := FALSE; END_IF;
END_REGION
END_FUNCTION_BLOCK

FUNCTION_BLOCK "Filling_Logic"   // FB2, LAD
{ S7_Optimized_Access := 'TRUE' }
VERSION : 0.1
   VAR_INPUT
      PS2_Filling_Station : Bool;
      FIC_B102 : Int;
      Liquid_AorB_in_Bottle_ml : Real;
      Liquid_AorB_pct : Int;
      PTRIG3 : Bool;
      PTRIG2 : Bool;
      Wait_to_fill : Time;
   END_VAR
   VAR_OUTPUT
      Outlet_of_tanks : Bool;
      Flow_ml_per_sec : Real;
      PTRIG1 : Bool;
      FillingData_LiqAorB_ml : Real;
   END_VAR
BEGIN

REGION Network 1
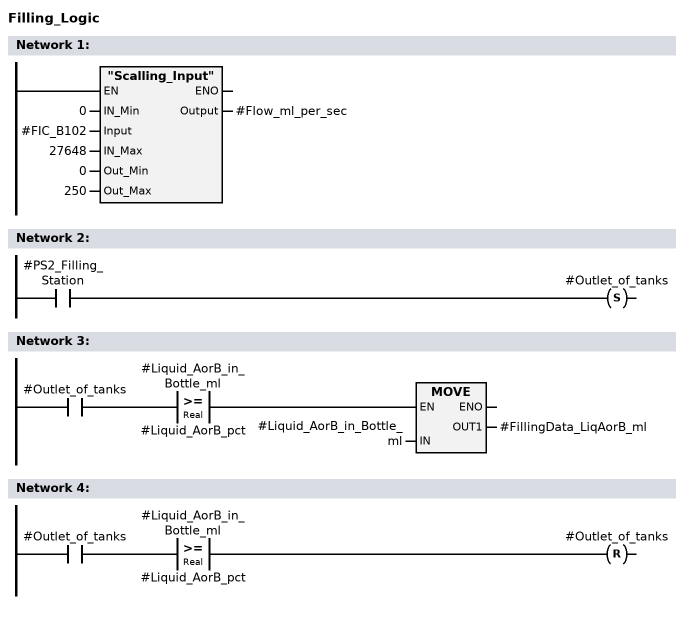
   RUNG wire#powerrail
      "Scalling_Input"(IN_Min := 0, Input := #FIC_B102, IN_Max := 27648, Out_Min := 0, Out_Max := 250, Output => #Flow_ml_per_sec)
   END_RUNG
   // the same network as SCL:
   "Scalling_Input"(IN_Min := 0,
                    Input := #FIC_B102,
                    IN_Max := 27648,
                    Out_Min := 0,
                    Out_Max := 250,
                    Output => #Flow_ml_per_sec);
END_REGION

REGION Network 2
   RUNG wire#powerrail
      Contact( #PS2_Filling_Station )
      S_Coil( #Outlet_of_tanks )
   END_RUNG
   // the same network as SCL:
   IF #PS2_Filling_Station THEN #Outlet_of_tanks := TRUE; END_IF;
END_REGION

REGION Network 3
   RUNG wire#powerrail
      Contact( #Outlet_of_tanks )
      { S7_Templates := "SrcType := Real" } GE_Contact(in1 := #Liquid_AorB_in_Bottle_ml, in2 := #Liquid_AorB_pct)
      Move(in := #Liquid_AorB_in_Bottle_ml, out1 => #FillingData_LiqAorB_ml)
   END_RUNG
   // the same network as SCL:
   IF #Outlet_of_tanks AND (#Liquid_AorB_in_Bottle_ml >= #Liquid_AorB_pct) THEN
       #FillingData_LiqAorB_ml := #Liquid_AorB_in_Bottle_ml;
   END_IF;
END_REGION

REGION Network 4
   RUNG wire#powerrail
      Contact( #Outlet_of_tanks )
      { S7_Templates := "SrcType := Real" } GE_Contact(in1 := #Liquid_AorB_in_Bottle_ml, in2 := #Liquid_AorB_pct)
      R_Coil( #Outlet_of_tanks )
   END_RUNG
   // the same network as SCL:
   IF #Outlet_of_tanks AND (#Liquid_AorB_in_Bottle_ml >= #Liquid_AorB_pct) THEN
       #Outlet_of_tanks := FALSE;
   END_IF;
END_REGION
END_FUNCTION_BLOCK

FUNCTION_BLOCK "Alarm_Logic"   // FB3, LAD
{ S7_Optimized_Access := 'TRUE' }
VERSION : 0.1
   VAR_TEMP   // added for the SCL form of the ladder/FBD networks
      _w1 : Bool;
      _w2 : Bool;
      _w3 : Bool;
      _w4 : Bool;
      _w5 : Bool;
      _w6 : Bool;
   END_VAR
BEGIN

REGION Network 1: Bottle Overfilled Alarm
   // 1. when total filled  liquid in the bottle is more than 100 ml, DECO block trigger the '1' bit of 'Alarm' word
   // 
   // for example: Normally    Alarm(Word) = 2#0000 0000 0000 0000
   // if filled  liquid in the bottle is more than 100 ml, Alarm(Word) = 2#0000 0000 0000 0010
   // 
   // 
   // all other alarms are programmed in the same way. Different bits of 'Alarm' word indicates different alarms.
   // 
   // This method is used, because with 'BOOL' variable Alarms can not be displayed on the HMI.
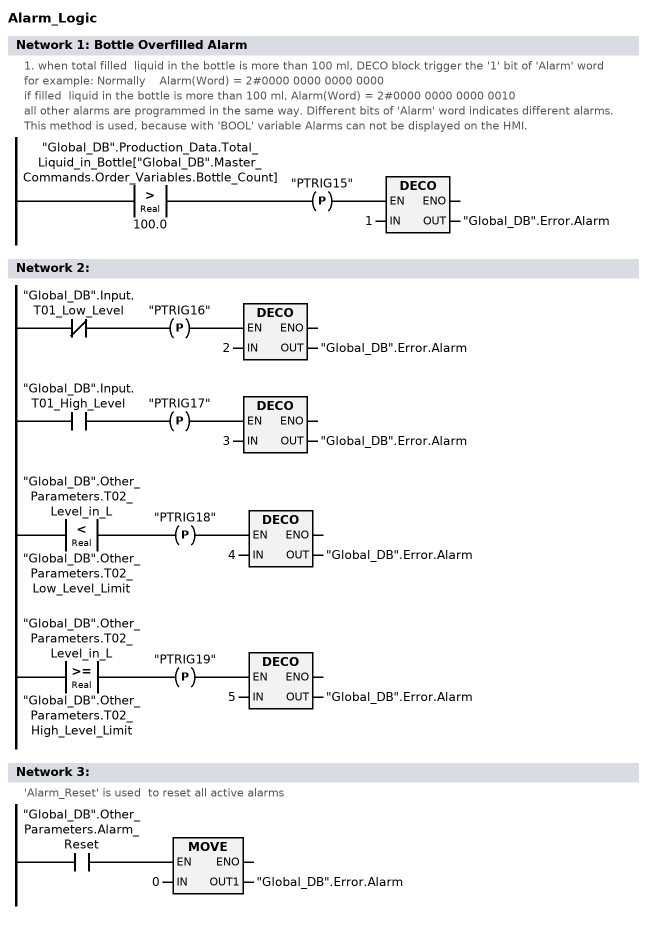
   #_w1 := "Global_DB".Production_Data.Total_Liquid_in_Bottle["Global_DB".Master_Commands.Order_Variables.Bottle_Count] > 100.0;
   #_w2 := #_w1 AND NOT "PTRIG15";   // rising edge
   "PTRIG15" := #_w1;
   IF #_w2 THEN "Global_DB".Error.Alarm := DECO(IN := 1); END_IF;
END_REGION

REGION Network 2
   #_w1 := NOT "Global_DB".Input.T01_Low_Level AND NOT "PTRIG16";   // rising edge
   "PTRIG16" := NOT "Global_DB".Input.T01_Low_Level;
   IF #_w1 THEN "Global_DB".Error.Alarm := DECO(IN := 2); END_IF;
   #_w2 := "Global_DB".Input.T01_High_Level AND NOT "PTRIG17";   // rising edge
   "PTRIG17" := "Global_DB".Input.T01_High_Level;
   IF #_w2 THEN "Global_DB".Error.Alarm := DECO(IN := 3); END_IF;
   #_w3 := "Global_DB".Other_Parameters.T02_Level_in_L < "Global_DB".Other_Parameters.T02_Low_Level_Limit;
   #_w4 := #_w3 AND NOT "PTRIG18";   // rising edge
   "PTRIG18" := #_w3;
   IF #_w4 THEN "Global_DB".Error.Alarm := DECO(IN := 4); END_IF;
   #_w5 := "Global_DB".Other_Parameters.T02_Level_in_L >= "Global_DB".Other_Parameters.T02_High_Level_Limit;
   #_w6 := #_w5 AND NOT "PTRIG19";   // rising edge
   "PTRIG19" := #_w5;
   IF #_w6 THEN "Global_DB".Error.Alarm := DECO(IN := 5); END_IF;
END_REGION

REGION Network 3
   // 'Alarm_Reset' is used  to reset all active alarms
   RUNG wire#powerrail
      Contact( "Global_DB".Other_Parameters.Alarm_Reset )
      Move(in := 0, out1 => "Global_DB".Error.Alarm)
   END_RUNG
   // the same network as SCL:
   IF "Global_DB".Other_Parameters.Alarm_Reset THEN "Global_DB".Error.Alarm := 0; END_IF;
END_REGION
END_FUNCTION_BLOCK

FUNCTION_BLOCK "Tank1"   // FB4, LAD
{ S7_Optimized_Access := 'TRUE' }
VERSION : 0.1
   VAR_INPUT
      EN_1 : Bool;
   END_VAR
   VAR_TEMP   // added for the SCL form of the ladder/FBD networks
      _w1 : Bool;
      _w2 : Bool;
      _w3 : Bool;
   END_VAR
BEGIN
